PopupScreen "Tank Status" 425x385
   Button "Button_1" at 365,1 size 56x38; TextOff 'Text'; PictureOff "Graphic_286"
      on Click: function_efd93a16("Tank Status", 0, 0, -1, -1, 1)
   Button "HmiScreenItemData_47" at 3,1 size 360x38; TextOn 'Back'; TextOff 'Automatic Ballast Tank Selection'
   Button "Button_4" at 14,64 size 100x23; TextOff 'FPT'; Authorization "Operate"
      on Press: function_b14e0dd5("504_Tank Grouping_DB2020_TANK ACTIV 1", 0)
      Appearance <- "504_Tank Grouping_DB2020_TANK ACTIV 1"
   Button "Button_2" at 338,151 size 79x32; TextOff '3'; Authorization "Operate"
      on Press: function_b14e0dd5("504_Tank Grouping_DB2020_GROUP ACTIV 3", 0)
      Appearance <- "504_Tank Grouping_DB2020_GROUP ACTIVE INT 3"
   Button "Button_3" at 338,185 size 79x32; TextOff '4'; Authorization "Operate"
      on Press: function_b14e0dd5("504_Tank Grouping_DB2020_GROUP ACTIV 4", 0)
      Appearance <- "504_Tank Grouping_DB2020_GROUP ACTIVE INT 4"
   Button "Button_10" at 339,219 size 79x32; TextOff '5'; Authorization "Operate"
      on Press: function_b14e0dd5("504_Tank Grouping_DB2020_GROUP ACTIV 5", 0)
      Appearance <- "504_Tank Grouping_DB2020_GROUP ACTIVE INT 5"
   Button "Button_11" at 339,253 size 79x32; TextOff '6'; Authorization "Operate"
      on Press: function_b14e0dd5("504_Tank Grouping_DB2020_GROUP ACTIV 6", 0)
      Appearance <- "504_Tank Grouping_DB2020_GROUP ACTIVE INT 6"
   Button "Button_12" at 339,288 size 79x32; TextOff '7'; Authorization "Operate"
      on Press: function_b14e0dd5("504_Tank Grouping_DB2020_GROUP ACTIV 7", 0)
      Appearance <- "504_Tank Grouping_DB2020_GROUP ACTIVE INT 7"
   Button "Button_7" at 338,83 size 79x32; TextOff '1'; Authorization "Operate"
      on Press: function_b14e0dd5("504_Tank Grouping_DB2020_GROUP ACTIV 1", 0)
      Appearance <- "504_Tank Grouping_DB2020_GROUP ACTIVE INT 1"
   Button "Button_8" at 338,117 size 79x32; TextOff '2'; Authorization "Operate"
      on Press: function_b14e0dd5("504_Tank Grouping_DB2020_GROUP ACTIV 2", 0)
      Appearance <- "504_Tank Grouping_DB2020_GROUP ACTIVE INT 2"
   Button "Button_9" at 14,96 size 100x23; TextOff 'TANK - 1P'; Authorization "Operate"
      on Press: function_b14e0dd5("504_Tank Grouping_DB2020_TANK ACTIV 2", 0)
      Appearance <- "504_Tank Grouping_DB2020_TANK ACTIV 2"
   Button "Button_14" at 14,128 size 100x23; TextOff 'TANK - 2P'; Authorization "Operate"
      on Press: function_b14e0dd5("504_Tank Grouping_DB2020_TANK ACTIV 4", 0)
      Appearance <- "504_Tank Grouping_DB2020_TANK ACTIV 4"
   Button "Button_15" at 14,160 size 100x23; TextOff 'TANK - 3P'; Authorization "Operate"
      on Press: function_b14e0dd5("504_Tank Grouping_DB2020_TANK ACTIV 6", 0)
      Appearance <- "504_Tank Grouping_DB2020_TANK ACTIV 6"
   Button "Button_16" at 14,193 size 100x23; TextOff 'TANK - 4P'; Authorization "Operate"
      on Press: function_b14e0dd5("504_Tank Grouping_DB2020_TANK ACTIV 8", 0)
      Appearance <- "504_Tank Grouping_DB2020_TANK ACTIV 8"
   Button "Button_17" at 14,225 size 100x23; TextOff 'TANK - 5P'; Authorization "Operate"
      on Press: function_b14e0dd5("504_Tank Grouping_DB2020_TANK ACTIV 10", 0)
      Appearance <- "504_Tank Grouping_DB2020_TANK ACTIV 10"
   Button "Button_18" at 14,257 size 100x23; TextOff 'TANK - 6P'; Authorization "Operate"
      on Press: function_b14e0dd5("504_Tank Grouping_DB2020_TANK ACTIV 12", 0)
      Appearance <- "504_Tank Grouping_DB2020_TANK ACTIV 12"
   Button "Button_19" at 14,290 size 100x23; TextOff 'TANK - APT'; Authorization "Operate"
      on Press: function_b14e0dd5("504_Tank Grouping_DB2020_TANK ACTIV 14", 0)
      Appearance <- "504_Tank Grouping_DB2020_TANK ACTIV 14"
   Button "Button_20" at 227,96 size 100x23; TextOff 'TANK - 1S'; Authorization "Operate"
      on Press: function_b14e0dd5("504_Tank Grouping_DB2020_TANK ACTIV 3", 0)
      Appearance <- "504_Tank Grouping_DB2020_TANK ACTIV 3"
   Button "Button_21" at 227,128 size 100x23; TextOff 'TANK - 2S'; Authorization "Operate"
      on Press: function_b14e0dd5("504_Tank Grouping_DB2020_TANK ACTIV 5", 0)
      Appearance <- "504_Tank Grouping_DB2020_TANK ACTIV 5"
   Button "Button_22" at 227,160 size 100x23; TextOff 'TANK - 3S'; Authorization "Operate"
      on Press: function_b14e0dd5("504_Tank Grouping_DB2020_TANK ACTIV 7", 0)
      Appearance <- "504_Tank Grouping_DB2020_TANK ACTIV 7"
   Button "Button_23" at 227,192 size 100x23; TextOff 'TANK - 4S'; Authorization "Operate"
      on Press: function_b14e0dd5("504_Tank Grouping_DB2020_TANK ACTIV 9", 0)
      Appearance <- "504_Tank Grouping_DB2020_TANK ACTIV 9"
   Button "Button_24" at 227,224 size 100x23; TextOff 'TANK - 5S'; Authorization "Operate"
      on Press: function_b14e0dd5("504_Tank Grouping_DB2020_TANK ACTIV 11", 0)
      Appearance <- "504_Tank Grouping_DB2020_TANK ACTIV 11"
   Button "Button_25" at 227,257 size 100x23; TextOff 'TANK - 6S'; Authorization "Operate"
      on Press: function_b14e0dd5("504_Tank Grouping_DB2020_TANK ACTIV 13", 0)
      Appearance <- "504_Tank Grouping_DB2020_TANK ACTIV 13"
   Switch "Switch_8" at 297,289 size 32x29; CaptionText 'Switch'; TextOn 'ON'; TextOff 'OFF'; Authorization "User administration"; PictureOff "Design_5_PilotLight_Green_Off"; PictureOn "Design_5_PilotLight_Green_On"
      on Change: InvertBit("80_From_HMI_Test Tank Request")
      Visibility <- "user_group"
      ProcessValue <- "504_Tank Grouping_DB2020_RUN"
   Circle "Circle_31" at 142,64 size 20x20
      Visibility <- "504_Tank Grouping_DB2020_RUN TANK 1"
      Appearance <- "504_Tank Grouping_DB2020_RUN TANK 1"
   Circle "Circle_4" at 121,130 size 20x20
      Appearance <- "504_Tank Grouping_DB2020_GROUP of TANK 4"
   Circle "Circle_6" at 120,161 size 20x20
      Appearance <- "504_Tank Grouping_DB2020_GROUP of TANK 6"
   Circle "Circle_7" at 120,98 size 20x20
      Appearance <- "504_Tank Grouping_DB2020_GROUP of TANK 2"
   Circle "Circle_8" at 120,226 size 20x20
      Appearance <- "504_Tank Grouping_DB2020_GROUP of TANK 10"
   Circle "Circle_10" at 120,194 size 20x20
      Appearance <- "504_Tank Grouping_DB2020_GROUP of TANK 8"
   Circle "Circle_11" at 120,291 size 20x20
      Appearance <- "504_Tank Grouping_DB2020_GROUP of TANK 14"
   Circle "Circle_12" at 120,258 size 20x20
      Appearance <- "504_Tank Grouping_DB2020_GROUP of TANK 12"
   IOField "I/O field_8" at 120,101 size 20x14; FormatPattern 99
      ProcessValue <- "504_Tank Grouping_DB2020_GROUP of TANK 2"
   IOField "I/O field_9" at 120,133 size 20x14; FormatPattern 99
      ProcessValue <- "504_Tank Grouping_DB2020_GROUP of TANK 4"
   IOField "I/O field_26" at 120,164 size 20x14; FormatPattern 99
      ProcessValue <- "504_Tank Grouping_DB2020_GROUP of TANK 6"
   IOField "I/O field_28" at 120,197 size 20x14; FormatPattern 99
      ProcessValue <- "504_Tank Grouping_DB2020_GROUP of TANK 8"
   IOField "I/O field_30" at 120,229 size 20x14; FormatPattern 99
      ProcessValue <- "504_Tank Grouping_DB2020_GROUP of TANK 10"
   IOField "I/O field_33" at 120,261 size 20x14; FormatPattern 99
      ProcessValue <- "504_Tank Grouping_DB2020_GROUP of TANK 12"
   IOField "I/O field_35" at 120,294 size 20x14; FormatPattern 99
      ProcessValue <- "504_Tank Grouping_DB2020_GROUP of TANK 14"
   Circle "Circle_13" at 199,130 size 20x20
      Appearance <- "504_Tank Grouping_DB2020_GROUP of TANK 5"
   Circle "Circle_14" at 199,160 size 20x20
      Appearance <- "504_Tank Grouping_DB2020_GROUP of TANK 7"
   Circle "Circle_15" at 199,98 size 20x20
      Appearance <- "504_Tank Grouping_DB2020_GROUP of TANK 3"
   Circle "Circle_16" at 199,225 size 20x20
      Appearance <- "504_Tank Grouping_DB2020_GROUP of TANK 11"
   Circle "Circle_17" at 199,193 size 20x20
      Appearance <- "504_Tank Grouping_DB2020_GROUP of TANK 9"
   Circle "Circle_18" at 199,258 size 20x20
      Appearance <- "504_Tank Grouping_DB2020_GROUP of TANK 13"
   IOField "I/O field_23" at 199,101 size 20x14; FormatPattern 99
      ProcessValue <- "504_Tank Grouping_DB2020_GROUP of TANK 3"
   IOField "I/O field_24" at 199,133 size 20x14; FormatPattern 99
      ProcessValue <- "504_Tank Grouping_DB2020_GROUP of TANK 5"
   IOField "I/O field_27" at 199,163 size 20x14; FormatPattern 99
      ProcessValue <- "504_Tank Grouping_DB2020_GROUP of TANK 7"
   IOField "I/O field_29" at 199,196 size 20x14; FormatPattern 99
      ProcessValue <- "504_Tank Grouping_DB2020_GROUP of TANK 9"
   IOField "I/O field_32" at 199,228 size 20x14; FormatPattern 99
      ProcessValue <- "504_Tank Grouping_DB2020_GROUP of TANK 11"
   IOField "I/O field_34" at 199,261 size 20x14; FormatPattern 99
      ProcessValue <- "504_Tank Grouping_DB2020_GROUP of TANK 13"
   Circle "Circle_32" at 142,97 size 20x20
      Visibility <- "504_Tank Grouping_DB2020_RUN TANK 2"
      Appearance <- "504_Tank Grouping_DB2020_RUN TANK 2"
   Circle "Circle_33" at 177,97 size 20x20
      Visibility <- "504_Tank Grouping_DB2020_RUN TANK 3"
      Appearance <- "504_Tank Grouping_DB2020_RUN TANK 3"
   Circle "Circle_34" at 142,129 size 20x20
      Visibility <- "504_Tank Grouping_DB2020_RUN TANK 4"
      Appearance <- "504_Tank Grouping_DB2020_RUN TANK 4"
   Circle "Circle_35" at 177,129 size 20x20
      Visibility <- "504_Tank Grouping_DB2020_RUN TANK 5"
      Appearance <- "504_Tank Grouping_DB2020_RUN TANK 5"
   Circle "Circle_36" at 142,161 size 20x20
      Visibility <- "504_Tank Grouping_DB2020_RUN TANK 6"
      Appearance <- "504_Tank Grouping_DB2020_RUN TANK 6"
   Circle "Circle_37" at 177,161 size 20x20
      Visibility <- "504_Tank Grouping_DB2020_RUN TANK 7"
      Appearance <- "504_Tank Grouping_DB2020_RUN TANK 7"
   Circle "Circle_38" at 142,193 size 20x20
      Visibility <- "504_Tank Grouping_DB2020_RUN TANK 8"
      Appearance <- "504_Tank Grouping_DB2020_RUN TANK 8"
   Circle "Circle_39" at 177,193 size 20x20
      Visibility <- "504_Tank Grouping_DB2020_RUN TANK 9"
      Appearance <- "504_Tank Grouping_DB2020_RUN TANK 9"
   Circle "Circle_40" at 142,225 size 20x20
      Visibility <- "504_Tank Grouping_DB2020_RUN TANK 10"
      Appearance <- "504_Tank Grouping_DB2020_RUN TANK 10"
   Circle "Circle_41" at 177,225 size 20x20
      Visibility <- "504_Tank Grouping_DB2020_RUN TANK 11"
      Appearance <- "504_Tank Grouping_DB2020_RUN TANK 11"
   Circle "Circle_42" at 142,258 size 20x20
      Visibility <- "504_Tank Grouping_DB2020_RUN TANK 12"
      Appearance <- "504_Tank Grouping_DB2020_RUN TANK 12"
   Circle "Circle_43" at 177,258 size 20x20
      Visibility <- "504_Tank Grouping_DB2020_RUN TANK 13"
      Appearance <- "504_Tank Grouping_DB2020_RUN TANK 13"
   Circle "Circle_44" at 142,290 size 20x20
      Visibility <- "504_Tank Grouping_DB2020_RUN TANK 14"
      Appearance <- "504_Tank Grouping_DB2020_RUN TANK 14"
   TextField "Text field_7" at 169,297 size 136x18; Text 'Test Tank Request'
      Visibility <- "user_group"
   Rectangle "Rectangle_6" at 337,45 size 82x37
      Visibility <- "504_Tank Grouping_DB2020_SetGroupSR"
   Button "Button_13" at 340,48 size 76x31; TextOff 'Set Group'; Authorization "Parameter Change"
      on Press: function_b14e0dd5("504_Tank Grouping_DB2020_SetGroup", 0)
      Appearance <- "504_Tank Grouping_DB2020_GROUP SET"
   Circle "Circle_5" at 120,64 size 20x20
      Appearance <- "504_Tank Grouping_DB2020_GROUP of TANK 1"
   IOField "I/O field_7" at 120,67 size 20x14; FormatPattern 99
      ProcessValue <- "504_Tank Grouping_DB2020_GROUP of TANK 1"
   Button "Button_6" at 82,331 size 256x47; TextOff 'Text'; Authorization "Operate"; PictureList "Water Level Override"
      on Press: function_b14e0dd5("2062_Warning_Data_Water Level Override", 0)
      ProcessValue <- "2062_Warning_Data_Water Level Override_Aux"

PopupScreen "IGG Start Confirm" 600x385
   Button "Button_1" at 554,1 size 42x31; TextOff 'Text'; PictureOff "Graphic_286"
      on Click: function_efd93a16("IGG Start Confirm", 0, 0, -1, -1, 1)
   Button "HmiScreenItemData_47" at 3,1 size 550x31; TextOn 'Back'; TextOff 'Inert Gas Generator Process Start Confirm'
   Button "HmiScreenItemData_4" at 308,265 size 212x66; TextOn 'CANCEL'; TextOff 'Cancel'; Authorization "Operate"
      on Release: function_efd93a16("IGG Start Confirm", 300, 200, -1, -1, 1)
   TextField "Text field_1" at 34,49 size 534x184; Text 'Acknowledging This The Inert Gas Generator Process Will Start. Machinery may start unexpectedly. Wear Personal Protection Equipment and Ear Defenders in The IGG Room.'
   TextField "Text field_2" at 163,220 size 300x46; Text 'ARE YOU SURE?'
   Button "HmiScreenItemData_1" at 86,275 size 169x47; TextOn 'START'; TextOff 'Start'; Authorization "Operate"
      on Press: function_b14e0dd5("80_From_HMI_RUN_IGG", 0); ResetBit("80_From_HMI_STOP_IGG")
      ObjectEnable <- "82_To_HMI_CRNT_MODE_IGG"
      on Release: function_efd93a16("IGG Start Confirm", 300, 200, -1, -1, 1)

PopupScreen "IGG Stop Confirm" 600x385
   Button "Button_1" at 554,1 size 42x31; TextOff 'Text'; PictureOff "Graphic_286"
      on Click: function_efd93a16("IGG Stop Confirm", 0, 0, -1, -1, 1)
   Button "HmiScreenItemData_47" at 3,1 size 550x31; TextOn 'Back'; TextOff 'Ballast Water Treatment Process Stop Confirm'
   Button "HmiScreenItemData_4" at 308,265 size 212x66; TextOn 'CANCEL'; TextOff 'Cancel'; Authorization "Operate"
      on Release: function_efd93a16("IGG Stop Confirm", 300, 200, -1, -1, 1)
   TextField "Text field_1" at 33,49 size 528x184; Text 'Acknowledging This The Inert Gas Generator Process Will Stop. Machinery may start unexpectedly. Wear Personal Protection Equipment and Ear Defenders in The IGG Room.'
   TextField "Text field_2" at 163,220 size 300x46; Text 'ARE YOU SURE?'
   Button "HmiScreenItemData_2" at 86,275 size 169x47; TextOn 'STOP'; TextOff 'Stop'; Authorization "Operate"
      on Press: ResetBit("80_From_HMI_RUN_IGG"); function_b14e0dd5("80_From_HMI_STOP_IGG", 0)
      ObjectEnable <- "82_To_HMI_CRNT_MODE_IGG"
      on Release: function_efd93a16("IGG Stop Confirm", 300, 200, -1, -1, 1)

PopupScreen "BWTS Start Confirm" 600x385
   Button "Button_1" at 554,1 size 42x31; TextOff 'Text'; PictureOff "Graphic_286"
      on Click: function_efd93a16("BWTS Start Confirm", 0, 0, -1, -1, 1)
   Button "HmiScreenItemData_47" at 3,1 size 550x31; TextOn 'Back'; TextOff 'Ballast Water Treatment Process Start Confirm'
   Button "HmiScreenItemData_4" at 308,265 size 212x66; TextOn 'CANCEL'; TextOff 'Cancel'; Authorization "Operate"
      on Release: function_efd93a16("BWTS Start Confirm", 0, 0, -1, -1, 1)
   Button "HmiScreenItemData_3" at 86,275 size 169x47; TextOn 'START'; TextOff 'Start'; Authorization "Operate"
      on Release: ActivateScreen("Inert Gas Generator Plant", 0); function_efd93a16("BWTS Start Confirm", 300, 200, -1, -1, 1)
      on Press: function_b14e0dd5("2110_BTCS_CNTRL_DB_START_SEQ", 0)
      ObjectEnable <- "82_To_HMI_CRNT_MODE_GCU"
   TextField "Text field_1" at 3,49 size 594x184; Text 'Acknowledging This The Ballast Water Treatment Process Will Start. Machines may start unexpectedly. Wear Personal Protection Equipment and Ear Defenders in The IGG Room.'
   TextField "Text field_2" at 163,220 size 300x46; Text 'ARE YOU SURE?'

PopupScreen "BWTS Stop Confirm" 600x385
   Button "Button_1" at 554,1 size 42x31; TextOff 'Text'; PictureOff "Graphic_286"
      on Click: function_efd93a16("BWTS Stop Confirm", 0, 0, -1, -1, 1)
   Button "HmiScreenItemData_47" at 3,1 size 550x31; TextOn 'Back'; TextOff 'Ballast Water Treatment Process Stop Confirm'
   Button "HmiScreenItemData_4" at 308,265 size 212x66; TextOn 'CANCEL'; TextOff 'Cancel'; Authorization "Operate"
      on Release: function_efd93a16("BWTS Stop Confirm", 0, 0, -1, -1, 1)
   TextField "Text field_1" at 3,49 size 588x184; Text 'Acknowledging This The Ballast Water Treatment Process Will Stop. Machines may start unexpectedly. Wear Personal Protection Equipment and Ear Defenders in The IGG Room.'
   TextField "Text field_2" at 163,220 size 300x46; Text 'ARE YOU SURE?'
   Button "HmiScreenItemData_1" at 86,275 size 169x47; TextOn 'STOP'; TextOff 'Stop'; Authorization "Operate"
      on Release: function_efd93a16("BWTS Stop Confirm", 300, 200, -1, -1, 1)
      on Press: function_b14e0dd5("2110_BTCS_CNTRL_DB_STOP_SEQ", 0)
      ObjectEnable <- "82_To_HMI_CRNT_MODE_GCU"

PopupScreen "Lost Comunication" 700x600
   GraphicView "Graphic view_4" at 0,0 size 700x600; Picture "Graphic_298"
   Button "Button_1" at 0,0 size 700x596; TextOff 'Communication Lost'

PopupScreen "CV 405 Grafics" 810x675
   Button "Button_1" at 753,0 size 56x40; TextOff 'Text'; PictureOff "Graphic_286"
      on Click: function_efd93a16("CV 405 Grafics", 0, 0, -1, -1, 1)
   GraphicView "Graphic view_2" at 2,2 size 751x35; Picture "Graphic_287"
   TextField "Text field_1" at 248,7 size 327x26; Text 'PGC IG PRESSURE MODULATION'
   TrendView "Trend view_2" at 1,39 size 809x635
      ValueAxis2End <- "84_Setpoints_PIT416_HighHigh"

PopupScreen "PGC Temperature Trends" 810x675
   on GenerateScreen: "TitleUpdater"()
   Button "Button_1" at 753,0 size 56x38; TextOff 'Text'; PictureOff "Graphic_286"
      on Click: function_efd93a16("PGC Temperature Trends", 0, 0, -1, -1, 1)
   GraphicView "Graphic view_2" at 2,2 size 751x35; Picture "Graphic_287"
   TrendView "Trend view_1" at 1,40 size 805x635
      Visibility <- "80_From_HMI_BWT_BYPASS"
   TextField "Text field_1" at 282,7 size 254x26; Text 'PGC Temperature Trends'

PopupScreen "PGC Setpoint Protection" 600x400
   TextField "Text field_2" at 73,293 size 178x22; Text 'PIT416 GAS TO DECK PRESSURE'
   IOField "I/O field_1" at 261,293 size 70x22; FormatPattern 9.9; Unit  Barg
      ProcessValue <- "12_AI_Data_PIT_416_SCALED"
   TextField "Text field_6" at 13,293 size 53x22; Text 'IW810'
   Button "Button_1" at 550,1 size 47x30; TextOff 'Text'; PictureOff "Graphic_286"
      on Click: function_efd93a16("PGC Setpoint Protection", 0, 0, -1, -1, 1)
   Button "HmiScreenItemData_47" at 3,1 size 546x30; TextOn 'Back'; TextOff 'Automatic PGC Setpoint Protection'
   TextField "Text field_29" at 337,216 size 75x22; Text 'Target'
   TextField "Text field_5" at 408,216 size 91x22; Text 'Safe Target'
   TextField "Text field_8" at 76,239 size 229x18; Text 'PIT416 GAS TO DECK PRESSURE'
   TextField "Text field_15" at 315,64 size 209x18; Text 'Activate Temperature Protection'
      Visibility <- "user_group"
   TextField "Text field_1" at 315,113 size 209x18; Text 'Activate Pressure Protection'
      Visibility <- "user_group"
   TextField "Text field_3" at 315,161 size 209x18; Text 'Activate Tank Change Protection'
      Visibility <- "user_group"
   TextField "Text field_23" at 73,326 size 178x22; Text 'E400 PT002 PGC PRESS'
   IOField "I/O field_46" at 261,326 size 70x22; FormatPattern s9.9; Unit  Barg
      ProcessValue <- "12_AI_Data_E_400_PT002_SCALED"
   TextField "Text field_24" at 13,326 size 53x22; Text 'IW818'
   TextField "Text field_51" at 73,360 size 178x22; Text 'E400 TT002 PGC TEMP'
   IOField "I/O field_101" at 261,360 size 70x22; FormatPattern s999; Unit  °C
      ProcessValue <- "12_AI_Data_E_400_TE002_SCALED"
   TextField "Text field_56" at 13,360 size 53x22; Text 'IW820'
   IOField "I/O field_62" at 528,326 size 60x22; Authorization "Parameter Change"; FormatPattern 9.9
      ProcessValue <- "84_Setpoints_E400_PT002_HighHigh"
   IOField "I/O field_61" at 464,326 size 60x22; Authorization "Parameter Change"; FormatPattern 9.9
      ProcessValue <- "84_Setpoints_E400_PT002_High"
   IOField "I/O field_66" at 464,360 size 60x22; Authorization "Parameter Change"; FormatPattern 999
      ProcessValue <- "84_Setpoints_E400_TT002_High"
   IOField "I/O field_67" at 528,360 size 60x22; Authorization "Parameter Change"; FormatPattern 999
      ProcessValue <- "84_Setpoints_E400_TT002_HighHigh"
   TextField "Text field_4" at 468,271 size 53x22; Text 'High'
   TextField "Text field_7" at 517,271 size 80x22; Text 'High High'
   IOField "I/O field_69" at 338,293 size 60x22; Authorization "Parameter Change"; FormatPattern 9.9
      ProcessValue <- "84_Setpoints_PIT416_LowLow"
   IOField "I/O field_70" at 401,293 size 60x22; Authorization "Parameter Change"; FormatPattern 9.9
      ProcessValue <- "84_Setpoints_PIT416_Low"
   IOField "I/O field_71" at 464,293 size 60x22; Authorization "Parameter Change"; FormatPattern 9.9
      ProcessValue <- "84_Setpoints_PIT416_High"
   IOField "I/O field_72" at 528,293 size 60x22; Authorization "Parameter Change"; FormatPattern 9.9
      ProcessValue <- "84_Setpoints_PIT416_HighHigh"
   TextField "Text field_9" at 340,272 size 60x22; Text 'Low Low'
   TextField "Text field_10" at 390,272 size 80x22; Text 'Low'
   TextField "Text field_11" at 16,63 size 166x18; Text 'Temperature Tolerance'
   TextField "Text field_12" at 16,97 size 137x18; Text 'Pressure Tolerance'
   TextField "Text field_13" at 16,132 size 110x18; Text 'Debounce time'
   IOField "I/O field_5" at 218,128 size 65x28; Authorization "Commissioning"; FormatPattern 999; Unit s
      ProcessValue <- "84_Setpoints_Tank Close TimeOut"
   Button "Button_2" at 210,163 size 78x31; TextOn 'RESET'; TextOff 'Reset'; Authorization "Operate"
      on Press: function_b14e0dd5("Setpoint Override_DB_Reset", 0)
      Appearance <- "Setpoint Override_DB_Set Pressure"
   IOField "I/O field_6" at 218,93 size 65x28; Authorization "Commissioning"; FormatPattern 9.99; Unit Barg
      ProcessValue <- "84_Setpoints_E-400 PT002 Tolerance"
   IOField "I/O field_3" at 218,59 size 65x28; Authorization "Commissioning"; FormatPattern 999; Unit  °C
      ProcessValue <- "84_Setpoints_E-400 TT002 Tolerance"
   Switch "Switch_4" at 541,152 size 45x43; CaptionText 'Switch'; TextOff 'OFF'; TextOn 'pilot'; PictureOn "Design_5_PilotLight_Green_On"; PictureOff "Design_5_PilotLight_Green_Off"; Authorization "Commissioning"
      ProcessValue <- "80_From_HMI_Tank Close Protection"
      on Change: InvertBit("80_From_HMI_Tank Close Protection")
   TextField "Text field_14" at 241,214 size 46x25; Text 'Text'
   Switch "Switch_3" at 541,101 size 45x43; CaptionText 'Switch'; TextOff 'OFF'; TextOn 'pilot'; Authorization "Commissioning"; PictureOff "Design_5_PilotLight_Green_Off"; PictureOn "Design_5_PilotLight_Green_On"
      ProcessValue <- "80_From_HMI_PT002 Target Protection"
      on Change: InvertBit("80_From_HMI_PT002 Target Protection")
   Switch "Switch_2" at 541,49 size 45x43; CaptionText 'Switch'; TextOff 'OFF'; TextOn 'pilot'; Authorization "Commissioning"; PictureOff "Design_5_PilotLight_Green_Off"; PictureOn "Design_5_PilotLight_Green_On"
      on Change: InvertBit("80_From_HMI_TT002 Target Protection")
      ProcessValue <- "80_From_HMI_TT002 Target Protection"
   IOField "I/O field_2" at 337,235 size 75x28; Authorization "Commissioning"; FormatPattern 9.9; Unit Barg
      ProcessValue <- "84_Setpoints_PIT416_Target"
   IOField "I/O field_4" at 417,235 size 75x28; Authorization "Commissioning"; FormatPattern 9.9; Unit Barg
      ProcessValue <- "84_Setpoints_PIT416_Target_Safe"

PopupScreen "PGC Protection Warning" 665x250
   Button "Button_1" at 0,0 size 665x250; TextOff 'THE INERT GAS PRESSURE WAS AUTOMATICALY LIMITED TO PREVENT PROCESS GAS COMPRESOR OVERHEATING'; Authorization "Operating Mode"
      on Release: function_efd93a16("PGC Protection Warning", 0, 0, -1, -1, 1)
   Button "Button_2" at 208,187 size 250x35; TextOff 'CHECK SETTINGS'
      on Release: function_efd93a16("PGC Protection Warning", 0, 0, -1, -1, 1); function_efd93a16("PGC Setpoint Protection", 300, 200, -1, -1, 1)

PopupScreen "Start Treatment" 665x230
   Button "Button_1" at 0,0 size 665x230; TextOff 'Text'
   Button "Button_2" at 232,146 size 200x55; TextOff 'OK'; Authorization "Operate"
      on Release: function_efd93a16("Start Treatment", 0, 0, -1, -1, 1); ActivateScreen("Inert Gas Generator Plant", 0)
   TextField "Text field_1" at 72,23 size 520x52; Text 'Treatment now required'
   TextField "Text field_2" at 16,73 size 644x64; Text 'Please Make Sure the Energy and Water Supply are Present and Sufficient'

PopupScreen "Start GCU for Re-Ox" 665x250
   Button "Button_1" at 0,0 size 665x250; TextOff 'Text'
   Button "Button_2" at 232,179 size 200x55; TextOff 'CONFIRM'; Authorization "Operate"
      on Release: function_efd93a16("Start GCU for Re-Ox", 0, 0, -1, -1, 1); ActivateScreen("Inert Gas Conditioning Plant", 0)
      on Press: function_b14e0dd5("80_From_HMI_GCU Start Confirmed", 0)
   TextField "Text field_1" at 8,6 size 647x100; Text 'Instalation Start Confirmation Required for Re-Ox Stage'
   TextField "Text field_2" at 16,109 size 644x64; Text 'Please Make Sure the Energy and Water Supply are Present and Sufficient'

PopupScreen "Time Until GCU Start Required" 750x270
   Button "Button_1" at 0,0 size 750x268; TextOff 'Text'
   Button "Button_2" at 269,198 size 200x55; TextOff 'OK'; Authorization "Operate"
      on Release: function_efd93a16("Time Until GCU Start Required", 0, 0, -1, -1, 1); ActivateScreen("Inert Gas Conditioning Plant", 0)
   TextField "Text field_1" at 5,4 size 726x133; Text 'Instalation Start Confirmation Required in hours and minutes for Re-Ox Stage'
   TextField "Text field_2" at 57,132 size 644x64; Text 'Please Make Sure the Energy and Water Supply are Present and Sufficient'
   IOField "I/O field_1" at 234,45 size 104x52; FormatPattern 99
      ProcessValue <- "Sequence Times_DB_Dwell Timer_Hours Left"
   IOField "I/O field_2" at 481,45 size 104x52; FormatPattern 99
      ProcessValue <- "Sequence Times_DB_Dwell Timer_Minutes Left"

PopupScreen "Time Until Treatment Required" 750x270
   Button "Button_1" at 0,0 size 750x270; TextOff 'Text'
   Button "Button_2" at 268,157 size 200x55; TextOff 'OK'; Authorization "Operate"
      on Click: function_efd93a16("Time Until Treatment Required", 0, 0, -1, -1, 1); ActivateScreen("Inert Gas Generator Plant", 0)
   TextField "Text field_1" at 6,24 size 728x100; Text 'Treatment required to start in hours and minutes'
   IOField "I/O field_1" at 207,72 size 104x52; FormatPattern 99
      ProcessValue <- "Sequence Times_DB_Pre-Dwell Timer_Hours Left"
   IOField "I/O field_2" at 470,72 size 104x52; FormatPattern 99
      ProcessValue <- "Sequence Times_DB_Pre-Dwell Timer_Minutes Left"

PopupScreen "Tank Times" 425x550
   TextField "Text field_34" at 35,501 size 206x35; Text 'TIMES VALID'
      Visibility <- "2102_TIME_CALCS_DB_TIMES_VALID"
   TextField "Text field_4" at 18,500 size 235x37; Text 'TIMES INVALID'
      Visibility <- "2102_TIME_CALCS_DB_TIMES_VALID"
   Button "HmiScreenItemData_47" at 4,1 size 359x38; TextOn 'Back'; TextOff 'Ballast Tank Durations'
   TextField "Text field_1" at 5,437 size 414x52; Text 'Did You Set Voyage Duration and Treatment Duration?'
   Button "HmiScreenItemData_14" at 4,40 size 416x27; TextOn 'Back'; TextOff 'Treatment Durations'
   TextField "Text field_14" at 13,80 size 85x18; Text 'Description'
   TextField "Text field_17" at 230,80 size 67x18; Text 'Setpoint'
   IOField "I/O field_10" at 216,118 size 92x27; Authorization "Operating Mode"; FormatPattern 999.99; Unit  Days
      ProcessValue <- "2115_VOYAGE_TIME_DAYS_VOYAGE_DAYS"
   IOField "I/O field_12" at 216,253 size 79x28; Authorization "Commissioning"; FormatPattern 999; Unit  Hrs
      ProcessValue <- "2110_BTCS_CNTRL_DB_DE_OX_HRS"
   IOField "I/O field_13" at 216,321 size 79x28; Authorization "Commissioning"; FormatPattern 999; Unit  Hrs
      ProcessValue <- "2110_BTCS_CNTRL_DB_DWELL_HRS"
   IOField "I/O field_14" at 216,355 size 79x28; Authorization "Commissioning"; FormatPattern 999; Unit  Hrs
      ProcessValue <- "2110_BTCS_CNTRL_DB_RE_OX_HRS"
   IOField "I/O field_15" at 216,389 size 79x28; Authorization "Commissioning"; FormatPattern 999; Unit  Hrs
      ProcessValue <- "2110_BTCS_CNTRL_DB_POST_DWELL_HRS"
   Button "HmiScreenItemData_11" at 12,114 size 203x35; TextOn 'Back'; TextOff 'Voyage A'
   Button "HmiScreenItemData_12" at 12,219 size 203x28; TextOn 'Back'; TextOff 'Pre Dwell Time'
   Button "HmiScreenItemData_13" at 12,253 size 203x28; TextOn 'Back'; TextOff 'De-Oxygenation Minimum Time'
   Button "HmiScreenItemData_43" at 12,321 size 203x28; TextOn 'Back'; TextOff 'Dwell Time'
   Button "HmiScreenItemData_44" at 12,355 size 203x28; TextOn 'Back'; TextOff 'Re-Oxygenation Time'
   Button "HmiScreenItemData_45" at 12,389 size 203x28; TextOn 'Back'; TextOff 'Post Dwell Time'
   IOField "I/O field_17" at 236,155 size 79x28; Authorization "User administration"; FormatPattern 999; Unit  Hrs
      ProcessValue <- "2110_BTCS_CNTRL_DB_TOT_SEQ_HRS"
   Button "HmiScreenItemData_42" at 12,155 size 203x28; TextOn 'Back'; TextOff 'Total Treatment Time'
   TextField "Text field_11" at 355,80 size 36x18; Text 'ETA'
   IOField "I/O field_16" at 332,219 size 83x28; Authorization "User administration"; FormatPattern 999; Unit  min
      ProcessValue <- "2102_TIME_CALCS_DB_PRE_DWELL_MINS_RMNG"
   IOField "I/O field_18" at 332,253 size 83x28; Authorization "User administration"; FormatPattern 999; Unit  min
   IOField "I/O field_19" at 332,321 size 83x28; FormatPattern 999; Unit  min
      ProcessValue <- "2102_TIME_CALCS_DB_DWELL_MINS_RMNG"
   IOField "I/O field_20" at 332,355 size 83x28; FormatPattern 999; Unit  min
      ProcessValue <- "2102_TIME_CALCS_DB_RE_OX_MINS_RMNG"
   IOField "I/O field_21" at 332,389 size 83x28; FormatPattern 999; Unit  min
      ProcessValue <- "2102_TIME_CALCS_DB_POST_DWELL_MINS_RMNG"
   IOField "I/O field_22" at 332,155 size 83x28; Authorization "User administration"; FormatPattern 999; Unit  Hrs
      ProcessValue <- "2110_BTCS_CNTRL_DB_RMNG_SEQ_HRS"
   IOField "I/O field_1" at 216,287 size 79x28; Authorization "Commissioning"; FormatPattern 999; Unit  Hrs
      ProcessValue <- "2110_BTCS_CNTRL_DB_DE_OX_SP_HRS"
   Button "HmiScreenItemData_6" at 12,287 size 203x28; TextOn 'Back'; TextOff 'De-Oxygenation Setpoint Time'
   Button "HmiScreenItemData_7" at 332,71 size 83x35; TextOn 'CONTINUE'; TextOff 'Continue'; Authorization "Operating Mode"
      on Press: InvertBit("80_From_HMI_TIMER RST Supres")
      Appearance <- "80_From_HMI_TIMER RST Supres"
   IOField "I/O field_25" at 216,187 size 79x28; Authorization "User administration"; FormatPattern 999.9; Unit  min
      ProcessValue <- "504_Tank Grouping_DB2020_Sequence Time m Offset_Int"
   Button "HmiScreenItemData_2" at 12,187 size 203x28; TextOn 'Back'; TextOff 'Differential Treatment Time'
   IOField "I/O field_3" at 332,187 size 83x28; Authorization "User administration"; FormatPattern 999; Unit  min
      ProcessValue <- "504_Tank Grouping_DB2020_Diff Time Remain"
   IOField "I/O field_48" at 348,155 size 33x28; Authorization "User administration"; FormatPattern 99; Unit h
      ProcessValue <- "Sequence Times_DB_Treatment Timer_Hours Left"
   IOField "I/O field_51" at 316,155 size 33x28; Authorization "User administration"; FormatPattern 99; Unit d
      ProcessValue <- "Sequence Times_DB_Treatment Timer_Days Left"
   IOField "I/O field_52" at 380,155 size 35x28; Authorization "User administration"; FormatPattern 99; Unit m
      ProcessValue <- "Sequence Times_DB_Treatment Timer_Minutes Left"
   IOField "I/O field_43" at 332,187 size 83x28; Authorization "User administration"; FormatPattern 999; Unit  min
      ProcessValue <- "504_Tank Grouping_DB2020_Diff Time Remain"
   IOField "I/O field_44" at 380,219 size 35x28; Authorization "User administration"; FormatPattern 99; Unit m
      ProcessValue <- "Sequence Times_DB_Pre-Dwell Timer_Minutes Left"
   IOField "I/O field_45" at 348,219 size 33x28; Authorization "User administration"; FormatPattern 99; Unit h
      ProcessValue <- "Sequence Times_DB_Pre-Dwell Timer_Hours Left"
   IOField "I/O field_46" at 316,219 size 33x28; Authorization "User administration"; FormatPattern 99; Unit d
      ProcessValue <- "Sequence Times_DB_Pre-Dwell Timer_Days Left"
   IOField "I/O field_47" at 216,118 size 92x28; Authorization "Operating Mode"; FormatPattern 999.9; Unit  Days
      ProcessValue <- "Sequence Times_DB_Jurney Time"
   IOField "I/O field_49" at 248,155 size 33x28; Authorization "User administration"; FormatPattern 99; Unit h
      ProcessValue <- "Sequence Times_DB_Treatment Timer_Hours"
   IOField "I/O field_50" at 216,155 size 33x28; Authorization "User administration"; FormatPattern 99; Unit d
      ProcessValue <- "Sequence Times_DB_Treatment Timer_Days"
   IOField "I/O field_53" at 280,155 size 35x28; Authorization "User administration"; FormatPattern 99; Unit m
      ProcessValue <- "Sequence Times_DB_Treatment Timer_Minutes"
   IOField "I/O field_54" at 348,118 size 33x28; Authorization "User administration"; FormatPattern 99; Unit h
      ProcessValue <- "Sequence Times_DB_Jurney Timer_Hours Left"
   IOField "I/O field_55" at 309,118 size 40x28; Authorization "User administration"; FormatPattern 999; Unit d
      ProcessValue <- "Sequence Times_DB_Jurney Timer_Days Left"
   IOField "I/O field_56" at 380,118 size 35x28; Authorization "User administration"; FormatPattern 99; Unit m
      ProcessValue <- "Sequence Times_DB_Jurney Timer_Minutes Left"
   IOField "I/O field_57" at 216,219 size 79x28; Authorization "Commissioning"; FormatPattern 9999.9; Unit  Hrs
      ProcessValue <- "Sequence Times_DB_Pre-Dwell Time"
   IOField "I/O field_58" at 216,253 size 79x28; Authorization "Commissioning"; FormatPattern 999.9; Unit  Hrs
      ProcessValue <- "Sequence Times_DB_De-Ox Time"
   IOField "I/O field_59" at 380,253 size 35x28; Authorization "User administration"; FormatPattern 99; Unit m
      ProcessValue <- "Sequence Times_DB_De-Ox Timer_Minutes Left"
   IOField "I/O field_60" at 348,253 size 33x28; Authorization "User administration"; FormatPattern 99; Unit h
      ProcessValue <- "Sequence Times_DB_De-Ox Timer_Hours Left"
   IOField "I/O field_61" at 316,253 size 33x28; Authorization "User administration"; FormatPattern 99; Unit d
      ProcessValue <- "Sequence Times_DB_De-Ox Timer_Days Left"
   IOField "I/O field_62" at 216,287 size 79x28; Authorization "Commissioning"; FormatPattern 999.9; Unit  Hrs
      ProcessValue <- "Sequence Times_DB_De-Ox SP Time"
   IOField "I/O field_63" at 216,321 size 79x28; Authorization "Commissioning"; FormatPattern 999.9; Unit  Hrs
      ProcessValue <- "Sequence Times_DB_Dwell Time"
   IOField "I/O field_64" at 380,321 size 35x28; Authorization "User administration"; FormatPattern 99; Unit m
      ProcessValue <- "Sequence Times_DB_Dwell Timer_Minutes Left"
   IOField "I/O field_65" at 348,321 size 33x28; Authorization "User administration"; FormatPattern 99; Unit h
      ProcessValue <- "Sequence Times_DB_Dwell Timer_Hours Left"
   IOField "I/O field_66" at 316,321 size 33x28; Authorization "User administration"; FormatPattern 99; Unit d
      ProcessValue <- "Sequence Times_DB_Dwell Timer_Days Left"
   IOField "I/O field_2" at 216,355 size 79x28; Authorization "Commissioning"; FormatPattern 999.9; Unit  Hrs
      ProcessValue <- "Sequence Times_DB_Re-Ox Time"
   IOField "I/O field_67" at 380,355 size 35x28; Authorization "User administration"; FormatPattern 99; Unit m
      ProcessValue <- "Sequence Times_DB_Re-Ox Timer_Minutes Left"
   IOField "I/O field_68" at 348,355 size 33x28; Authorization "User administration"; FormatPattern 99; Unit h
      ProcessValue <- "Sequence Times_DB_Re-Ox Timer_Hours Left"
   IOField "I/O field_69" at 316,355 size 33x28; Authorization "User administration"; FormatPattern 99; Unit d
      ProcessValue <- "Sequence Times_DB_Re-Ox Timer_Days Left"
   IOField "I/O field_70" at 216,389 size 79x28; Authorization "Commissioning"; FormatPattern 999.9; Unit  Hrs
      ProcessValue <- "Sequence Times_DB_Post-Dwell Time"
   IOField "I/O field_71" at 380,389 size 35x28; Authorization "User administration"; FormatPattern 99; Unit m
      ProcessValue <- "Sequence Times_DB_Post-Dwell Timer_Minutes Left"
   IOField "I/O field_72" at 348,389 size 33x28; Authorization "User administration"; FormatPattern 99; Unit h
      ProcessValue <- "Sequence Times_DB_Post-Dwell Timer_Hours Left"
   IOField "I/O field_73" at 316,389 size 33x28; Authorization "User administration"; FormatPattern 99; Unit d
      ProcessValue <- "Sequence Times_DB_Post-Dwell Timer_Days Left"
   Button "HmiScreenItemData_1" at 263,499 size 116x39; TextOn 'ALL SET'; TextOff 'All Set'; Authorization "Commissioning"
      on Press: SetTag("2068_Sys_Status_Data_Times Visibil", 0)
      on Release: function_efd93a16("Tank Times", 300, 200, -1, -1, 1)
   Button "Button_1" at 364,1 size 56x38; TextOff 'Text'; PictureOff "Graphic_286"
      on Click: function_efd93a16("Tank Times", 300, 200, -1, -1, 1)
   Group "Group_1" at 18,500 size 235x37

PopupScreen "TANK Activ Warning" 665x250
   Button "Button_1" at 0,0 size 665x250; TextOff 'No TANK Selected. Select a TANK for Tank Treatment.'
      on Release: function_efd93a16("TANK Activ Warning", 300, 200, -1, -1, 1)
   Button "Button_2" at 208,187 size 250x35; TextOff 'OK, Select TANK'
      on Release: ActivateScreen("Balast Water Treatment Setup", 0); function_efd93a16("TANK Activ Warning", 0, 0, -1, -1, 1)

screen "Balast Water Treatment Plant Tank Pressure" 1280x800, template "Template"
   on GenerateScreen: "User_Change"(); "TitleUpdater"()
   Button "HmiScreenItemData_1" at 1,1 size 150x40; TextOn 'Back'; TextOff 'Main Index'
      on Release: ActivateScreen("02 Main Index", 0)
   TextField "Text field_63" at 383,107 size 72x30; Text 'Pre Dwell Time'
   Circle "Circle_29" at 1047,85 size 20x20
      Appearance <- "2102_TIME_CALCS_DB_POST_DWELL_TMR_DN"
   Button "HmiScreenItemData_9" at 10,60 size 158x27; TextOn 'Back'; TextOff 'BWTS Control'
   Button "HmiScreenItemData_4" at 14,150 size 75x47; TextOn 'Back'; TextOff 'Stop'; Authorization "Operate"
      on Release: function_efd93a16("BWTS Stop Confirm", 400, 200, -1, -1, 1)
      ObjectEnable <- "82_To_HMI_CRNT_MODE_GCU"
   Circle "Circle_20" at 137,105 size 29x29
      Appearance <- "80_From_HMI_RUN_IGG(1)"
   Button "HmiScreenItemData_3" at 14,93 size 75x47; TextOn 'Back'; TextOff 'Start'; Authorization "Operate"
      on Release: function_efd93a16("BWTS Start Confirm", 400, 200, -1, -1, 1)
      ObjectEnable <- "82_To_HMI_CRNT_MODE_GCU"
   Button "HmiScreenItemData_2" at 1129,1 size 150x40; TextOn 'Back'; TextOff 'BWTS Setup'
      on Release: ActivateScreen("Balast Water Treatment Setup", 0)
   TextField "Text field_1" at 290,107 size 68x30; Text 'Tank Selected'
   TextField "Text field_2" at 841,107 size 61x30; Text 'BWTS Started'
   TextField "Text field_3" at 568,107 size 62x30; Text 'IGGS Started'
   TextField "Text field_4" at 659,107 size 60x30; Text 'GCU Started'
   TextField "Text field_5" at 748,107 size 61x30; Text 'PGC Started'
   TextField "Text field_6" at 908,107 size 102x30; Text 'Gas Transfer Started'
   Circle "Circle_10" at 956,89 size 14x14
      Appearance <- "2110_BTCS_CNTRL_DB_BTCS_STEP"
   TextField "Text field_7" at 995,107 size 125x30; Text 'Treatment Cycle Completed'
   TextField "Text field_23" at 261,291 size 34x14; Text 'MBG'
   GraphicView "Graphic view_17" at 575,446 size 532x12; Picture "Graphic_151"
   Button "Button_13" at 252,437 size 37x30; TextOff 'DB&B'
   TextField "Text field_58" at 188,226 size 50x40; Text 'Safe Area'
   Button "Button_20" at 724,152 size 115x34; TextOff 'Re-Oxygenation'
      Appearance <- "2110_BTCS_CNTRL_DB_BTCS_STEP"
   Button "Button_21" at 845,152 size 93x34; TextOff 'Post Dwell'
      Appearance <- "2110_BTCS_CNTRL_DB_BTCS_STATE"
   Circle "Circle_1" at 137,105 size 29x29
      Appearance <- "2110_BTCS_CNTRL_DB_BTCS_STATE"
   Circle "Circle_8" at 775,89 size 14x14
      Appearance <- "2110_BTCS_CNTRL_DB_BTCS_STEP"
   Circle "Circle_9" at 685,89 size 14x14
      Appearance <- "100_GCU_AUTO_SEQ_DB_CRNT_STEP"
   Circle "Circle_11" at 595,89 size 14x14
      Appearance <- "51_SLAVE_STATUS_RUNNING"
   Circle "Circle_12" at 866,89 size 14x14
      Appearance <- "2110_BTCS_CNTRL_DB_BTCS_STEP"
   Circle "Circle_13" at 324,89 size 14x14
      Appearance <- "HMI Indication Logic_DB_Tank Selected"
   Circle "Circle_14" at 414,89 size 14x14
      Appearance <- "2102_TIME_CALCS_DB_PRE_DWELL_TMR_DN"
   Button "Button_3" at 626,152 size 93x34; TextOff 'Dwell'
      Appearance <- "2110_BTCS_CNTRL_DB_BTCS_STATE"
   Button "Button_5" at 944,152 size 93x34; TextOff 'Complete'
      Appearance <- "HMI Indication Logic_DB_Sequence Finished"
   TextField "Text field_61" at 202,107 size 71x30; Text 'FA Mode Selected'
   Circle "Circle_2" at 230,89 size 14x14
      Appearance <- "HMI Indication Logic_DB_FA Mode Selected"
   TextField "Text field_60" at 190,519 size 46x25; Text 'GCU'
   GraphicIOField "Graphic I/O field_4" at 187,543 size 53x55; PictureList "GCU"
      ProcessValue <- "100_GCU_AUTO_SEQ_DB_RNG"
   TextField "Text field_74" at 186,279 size 54x25; Text 'IGGS'
   GraphicIOField "Graphic I/O field_1" at 185,303 size 57x53; PictureList "IGGS"
      ProcessValue <- "14_DQ_Data_24PF1"
   TextField "Text field_62" at 183,359 size 60x20; Text 'Disabled'
   TextField "Text field_77" at 183,359 size 60x20; Text 'Enabled'
      Visibility <- "51_SLAVE_STATUS_RUNNING"
   Button "Button_8" at 178,280 size 70x105; TextOff 'Text'
      on Release: ActivateScreen("Inert Gas Generator Plant", 0)
   TextField "Text field_70" at 183,599 size 60x20; Text 'Disabled'
   TextField "Text field_71" at 183,599 size 60x20; Text 'Enabled'
      Visibility <- "100_GCU_AUTO_SEQ_DB_RNG"
   Button "Button_4" at 178,521 size 70x105; TextOff 'Text'
      on Release: ActivateScreen("Inert Gas Conditioning Plant", 0)
   GraphicIOField "Graphic I/O field_2" at 770,45 size 250x30; PictureList "Process time Banner"
      Visibility <- "2110_BTCS_CNTRL_DB_BTCS_STATE"
      ProcessValue <- "2110_BTCS_CNTRL_DB_BTCS_STATE"
   Button "Button_14" at 303,152 size 93x34; TextOff 'Unselected'
      Visibility <- "HMI Indication Logic_DB_Tank Selected"
      Appearance <- "HMI Indication Logic_DB_Tank Selected"
   Button "Button_15" at 404,152 size 93x34; TextOff 'Selected'
      Appearance <- "HMI Indication Logic_DB_Tank Selected"
   Button "Button_16" at 506,152 size 115x34; TextOff 'De-Oxygenation'
      Appearance <- "2110_BTCS_CNTRL_DB_BTCS_STEP"
   TextField "Text field_92" at 304,351 size 76x15; Text 'FIT-418-6P'
   TextField "Text field_98" at 304,308 size 76x15; Text 'FIT-420-6P'
   Button "HmiScreenItemData_19" at 1185,676 size 72x27; TextOn 'Back'; TextOff 'Status'
      on Press: function_efd93a16("Treatment Status", 100, 471, -1, 3, 1)
   Group "Group_6" at 298,44 size 241x30
   Circle "Circle_26" at 504,89 size 14x14
      Appearance <- "2102_TIME_CALCS_DB_Time_To_Treatment"
   TextField "Text field_134" at 470,107 size 75x30; Text 'Wait for IGGS Start'
   GraphicView "Graphic view_4" at 357,210 size 25x62; Picture "Graphic_183"
   GraphicView "Graphic view_5" at 265,210 size 25x62; Picture "Graphic_183"
   IOField "I/O field_31" at 1053,45 size 225x30; FormatPattern ???????????????
      ProcessValue <- "Current User"
   Button "HmiScreenItemData_8" at 772,732 size 503x40; TextOn 'Back'; TextOff 'Text'
   TextField "Screen title" at 783,728 size 496x50; Text 'Screen title'
   Bar "Bar_1" at 262,206 size 122x241; MinimumValue 0; MaximumValue 100
      ProcessValue <- "20_TANKS_IP_DATA_RIO_06_FIRST_TANK_TANKS_PRESS"
   Button "Button_48" at 273,396 size 100x25; TextOff 'DISABLED'
      on Release: function_efd93a16("Tank 6P Status", 168, 315, -1, 2, 1)
      Visibility <- "504_Tank Grouping_DB2020_GROUP of TANK 12"
   Circle "Circle_3" at 340,212 size 14x14
      Appearance <- "20_TANKS_IP_DATA_RIO_06_FIRST_TANK_BWT_LEVEL_HIHI"
   TextField "Text field_125" at 295,212 size 51x14; Text 'LS425-6P'
   Polyline "Polyline_1" at 261,205 size 123x240
      Visibility <- "504_Tank Grouping_DB2020_RUN TANK 12"
   TextField "Text field_64" at 288,273 size 74x20; Text 'Tank - 6P'
   Bar "Bar_2" at 394,206 size 122x241; MinimumValue 0; MaximumValue 100
      ProcessValue <- "20_TANKS_IP_DATA_RIO_05_FIRST_TANK_TANKS_PRESS"
   Button "Button_44" at 406,396 size 100x25; TextOff 'DISABLED'
      on Release: function_efd93a16("Tank 5P Status", 168, 315, -1, 2, 1)
      Visibility <- "504_Tank Grouping_DB2020_GROUP of TANK 10"
   Circle "Circle_4" at 472,212 size 14x14
      Appearance <- "20_TANKS_IP_DATA_RIO_05_FIRST_TANK_BWT_LEVEL_HIHI"
   TextField "Text field_124" at 427,212 size 51x14; Text 'LS425-5P'
   Polyline "Polyline_2" at 392,205 size 123x240
      Visibility <- "504_Tank Grouping_DB2020_RUN TANK 10"
   TextField "Text field_8" at 418,275 size 74x20; Text 'Tank - 5P'
   Bar "Bar_3" at 525,206 size 122x241; MinimumValue 0; MaximumValue 100
      ProcessValue <- "20_TANKS_IP_DATA_RIO_04_FIRST_TANK_TANKS_PRESS"
   Button "Button_40" at 537,395 size 100x25; TextOff 'DISABLED'
      on Release: function_efd93a16("Tank 4P Status", 168, 315, -1, 2, 1)
      Visibility <- "504_Tank Grouping_DB2020_GROUP of TANK 8"
   Circle "Circle_5" at 604,212 size 14x14
      Appearance <- "20_TANKS_IP_DATA_RIO_04_FIRST_TANK_BWT_LEVEL_HIHI"
   TextField "Text field_123" at 559,212 size 51x14; Text 'LS425-4P'
   Polyline "Polyline_3" at 525,205 size 123x240
      Visibility <- "504_Tank Grouping_DB2020_RUN TANK 8"
   TextField "Text field_9" at 553,275 size 74x20; Text 'Tank - 4P'
   Bar "Bar_4" at 657,206 size 122x241; MinimumValue 0; MaximumValue 100
      ProcessValue <- "20_TANKS_IP_DATA_RIO_03_FIRST_TANK_TANKS_PRESS"
   Button "Button_36" at 668,395 size 100x25; TextOff 'DISABLED'
      on Release: function_efd93a16("Tank 3P Status", 168, 315, -1, 0, 1)
      Visibility <- "504_Tank Grouping_DB2020_GROUP of TANK 6"
   Circle "Circle_7" at 736,212 size 14x14
      Appearance <- "20_TANKS_IP_DATA_RIO_03_FIRST_TANK_BWT_LEVEL_HIHI"
   TextField "Text field_122" at 691,212 size 51x14; Text 'LS425-3P'
   Polyline "Polyline_4" at 656,205 size 123x240
      Visibility <- "504_Tank Grouping_DB2020_RUN TANK 6"
   TextField "Text field_14" at 680,275 size 74x20; Text 'Tank - 3P'
   Bar "Bar_5" at 789,206 size 122x241; MinimumValue 0; MaximumValue 100
      ProcessValue <- "20_TANKS_IP_DATA_RIO_02_FIRST_TANK_TANKS_PRESS"
   Button "Button_32" at 802,396 size 100x25; TextOff 'DISABLED'
      on Release: function_efd93a16("Tank 2P Status", 168, 315, -1, 0, 1)
      Visibility <- "504_Tank Grouping_DB2020_GROUP of TANK 4"
   Circle "Circle_15" at 868,212 size 14x14
      Appearance <- "20_TANKS_IP_DATA_RIO_02_FIRST_TANK_BWT_LEVEL_HIHI"
   TextField "Text field_121" at 823,212 size 51x14; Text 'LS425-2P'
   Polyline "Polyline_5" at 789,205 size 123x240
      Visibility <- "504_Tank Grouping_DB2020_RUN TANK 4"
   TextField "Text field_15" at 816,275 size 74x20; Text 'Tank - 2P'
   Bar "Bar_6" at 922,205 size 122x241; MinimumValue 0; MaximumValue 100
      ProcessValue <- "20_TANKS_IP_DATA_RIO_01_FIRST_TANK_TANKS_PRESS"
   Button "Button_52" at 934,395 size 100x25; TextOff 'DISABLED'
      on Release: function_efd93a16("Tank 1P Status", 168, 315, -1, 0, 1)
      Visibility <- "504_Tank Grouping_DB2020_GROUP of TANK 2"
   Circle "Circle_16" at 999,211 size 14x14
      Appearance <- "20_TANKS_IP_DATA_RIO_01_SECOND_TANK_BWT_LEVEL_HIHI"
   TextField "Text field_120" at 955,211 size 51x14; Text 'LS425-1P'
   Polyline "Polyline_6" at 921,205 size 123x240
      Visibility <- "504_Tank Grouping_DB2020_RUN TANK 2"
   GraphicView "Graphic view_6" at 127,446 size 591x12; Picture "Graphic_151"
   TextField "Text field_16" at 947,275 size 74x20; Text 'Tank - 1P'
   Bar "Bar_7" at 1096,334 size 122x241; MinimumValue 0; MaximumValue 100
      ProcessValue <- "20_TANKS_IP_DATA_RIO_01_FIRST_TANK_TANKS_PRESS"
   Circle "Circle_24" at 1168,339 size 14x14
      Appearance <- "20_TANKS_IP_DATA_RIO_01_FIRST_TANK_BWT_LEVEL_HIHI"
   TextField "Text field_133" at 1139,339 size 35x14; Text 'LS425'
   Polyline "Polyline_14" at 1095,332 size 125x242
      Visibility <- "504_Tank Grouping_DB2020_RUN TANK 1"
   Button "Button_56" at 1110,524 size 100x25; TextOff 'DISABLED'
      on Release: function_efd93a16("Tank FP Status", 168, 315, -1, 0, 1)
      Visibility <- "504_Tank Grouping_DB2020_GROUP of TANK 1"
   TextField "Text field_17" at 1111,400 size 111x20; Text 'Fore PeakTank'
   Bar "Bar_8" at 922,458 size 122x258; MinimumValue 0; MaximumValue 100
      ProcessValue <- "20_TANKS_IP_DATA_RIO_01_FIRST_TANK_TANKS_PRESS"
   Button "Button_54" at 933,661 size 100x25; TextOff 'DISABLED'
      on Release: function_efd93a16("Tank 1S Status", 168, 315, -1, 0, 1)